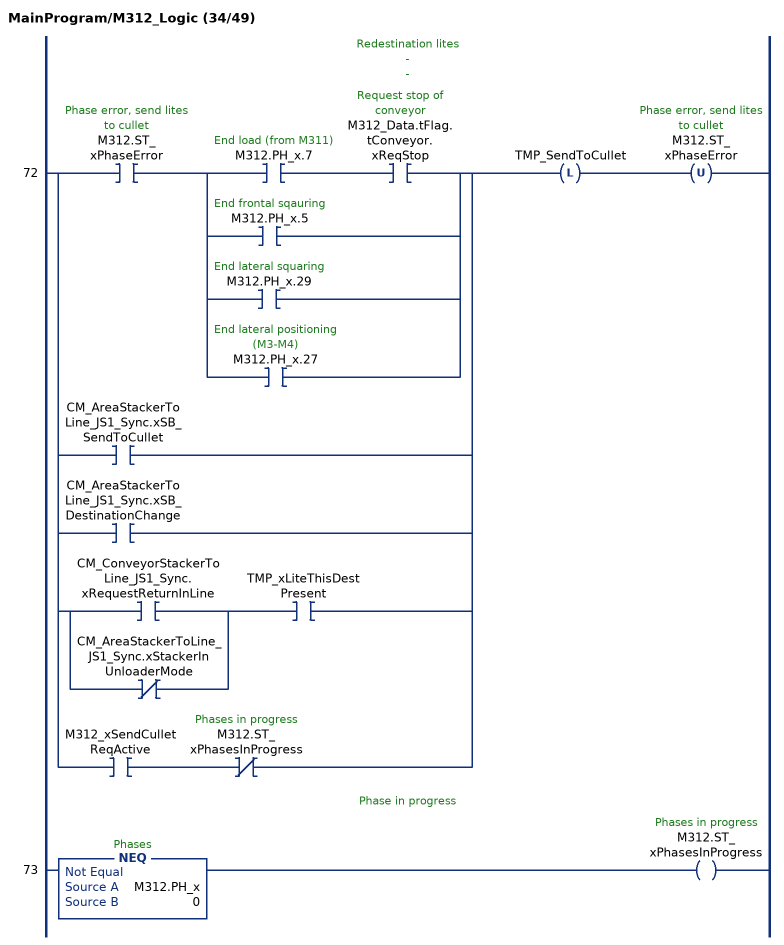
   // Redestination lites
   // -
   // -
   72: [XIC(M312.ST_xPhaseError) [XIC(M312.PH_x.7) XIC(M312_Data.tFlag.tConveyor.xReqStop) ,XIC(M312.PH_x.5) ,XIC(M312.PH_x.29) ,XIC(M312.PH_x.27) ] ,[XIC(CM_AreaStackerToLine_JS1_Sync.xSB_SendToCullet) ,XIC(CM_AreaStackerToLine_JS1_Sync.xSB_DestinationChange) ] ,[XIC(CM_ConveyorStackerToLine_JS1_Sync.xRequestReturnInLine) ,XIO(CM_AreaStackerToLine_JS1_Sync.xStackerInUnloaderMode) ] XIC(TMP_xLiteThisDestPresent) ,XIC(M312_xSendCulletReqActive) XIO(M312.ST_xPhasesInProgress) ]OTL(TMP_SendToCullet)OTU(M312.ST_xPhaseError);
   // Phase in progress
   73: NEQ(M312.PH_x,0)OTE(M312.ST_xPhasesInProgress);
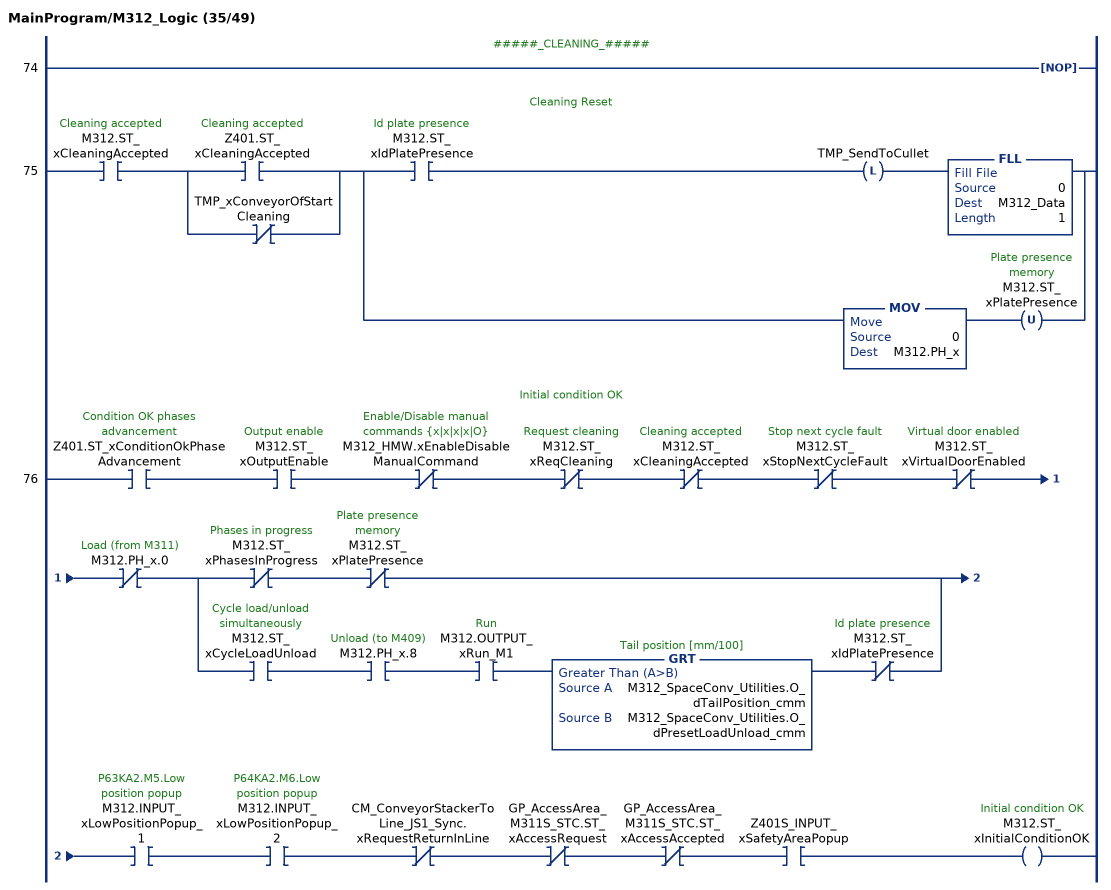
   // #####_CLEANING_#####
   74: NOP();
   // Cleaning Reset
   75: XIC(M312.ST_xCleaningAccepted)[XIC(Z401.ST_xCleaningAccepted) ,XIO(TMP_xConveyorOfStartCleaning) ][XIC(M312.ST_xIdPlatePresence) OTL(TMP_SendToCullet) FLL(0,M312_Data,1) ,MOV(0,M312.PH_x) OTU(M312.ST_xPlatePresence) ];
   // Initial condition OK
   76: XIC(Z401.ST_xConditionOkPhaseAdvancement)XIC(M312.ST_xOutputEnable)XIO(M312_HMW.xEnableDisableManualCommand)XIO(M312.ST_xReqCleaning)XIO(M312.ST_xCleaningAccepted)XIO(M312.ST_xStopNextCycleFault)XIO(M312.ST_xVirtualDoorEnabled)XIO(M312.PH_x.0)[XIO(M312.ST_xPhasesInProgress) XIO(M312.ST_xPlatePresence) ,XIC(M312.ST_xCycleLoadUnload) XIC(M312.PH_x.8) XIC(M312.OUTPUT_xRun_M1) GRT(M312_SpaceConv_Utilities.O_dTailPosition_cmm,M312_SpaceConv_Utilities.O_dPresetLoadUnload_cmm) XIO(M312.ST_xIdPlatePresence) ]XIC(M312.INPUT_xLowPositionPopup_1)XIC(M312.INPUT_xLowPositionPopup_2)XIO(CM_ConveyorStackerToLine_JS1_Sync.xRequestReturnInLine)XIO(GP_AccessArea_M311S_STC.ST_xAccessRequest)XIO(GP_AccessArea_M311S_STC.ST_xAccessAccepted)XIC(Z401S_INPUT_xSafetyAreaPopup)OTE(M312.ST_xInitialConditionOK);
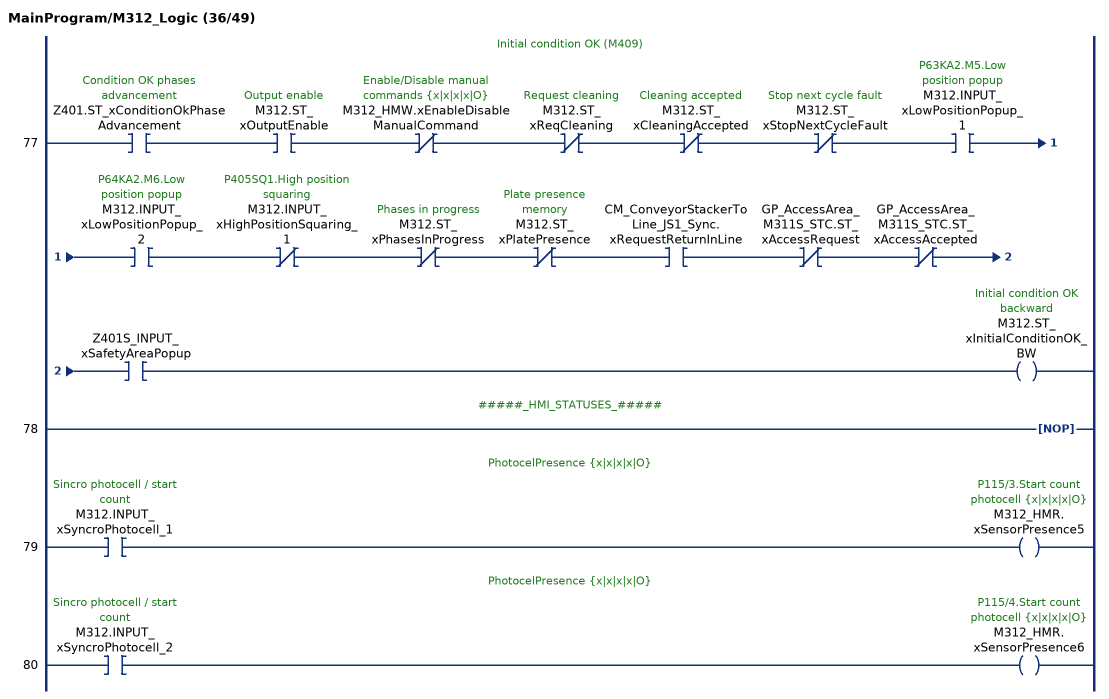
   // Initial condition OK (M409)
   77: XIC(Z401.ST_xConditionOkPhaseAdvancement)XIC(M312.ST_xOutputEnable)XIO(M312_HMW.xEnableDisableManualCommand)XIO(M312.ST_xReqCleaning)XIO(M312.ST_xCleaningAccepted)XIO(M312.ST_xStopNextCycleFault)XIC(M312.INPUT_xLowPositionPopup_1)XIC(M312.INPUT_xLowPositionPopup_2)XIO(M312.INPUT_xHighPositionSquaring_1)XIO(M312.ST_xPhasesInProgress)XIO(M312.ST_xPlatePresence)XIC(CM_ConveyorStackerToLine_JS1_Sync.xRequestReturnInLine)XIO(GP_AccessArea_M311S_STC.ST_xAccessRequest)XIO(GP_AccessArea_M311S_STC.ST_xAccessAccepted)XIC(Z401S_INPUT_xSafetyAreaPopup)OTE(M312.ST_xInitialConditionOK_BW);
   // #####_HMI_STATUSES_#####
   78: NOP();
   // PhotocelPresence {x|x|x|x|O}
   79: XIC(M312.INPUT_xSyncroPhotocell_1)OTE(M312_HMR.xSensorPresence5);
   // PhotocelPresence {x|x|x|x|O}
   80: XIC(M312.INPUT_xSyncroPhotocell_2)OTE(M312_HMR.xSensorPresence6);
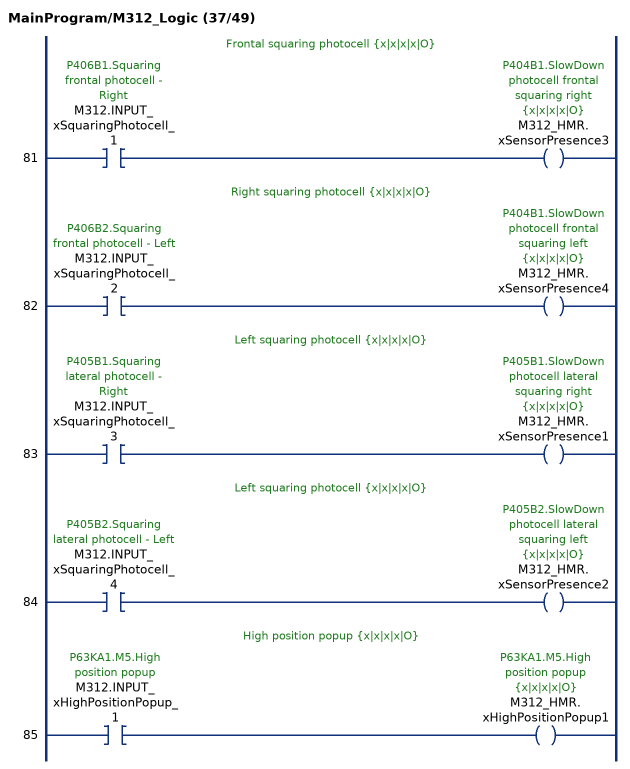
   // Frontal squaring photocell {x|x|x|x|O}
   81: XIC(M312.INPUT_xSquaringPhotocell_1)OTE(M312_HMR.xSensorPresence3);
   // Right squaring photocell {x|x|x|x|O}
   82: XIC(M312.INPUT_xSquaringPhotocell_2)OTE(M312_HMR.xSensorPresence4);
   // Left squaring photocell {x|x|x|x|O}
   83: XIC(M312.INPUT_xSquaringPhotocell_3)OTE(M312_HMR.xSensorPresence1);
   // Left squaring photocell {x|x|x|x|O}
   84: XIC(M312.INPUT_xSquaringPhotocell_4)OTE(M312_HMR.xSensorPresence2);
   // High position popup {x|x|x|x|O}
   85: XIC(M312.INPUT_xHighPositionPopup_1)OTE(M312_HMR.xHighPositionPopup1);
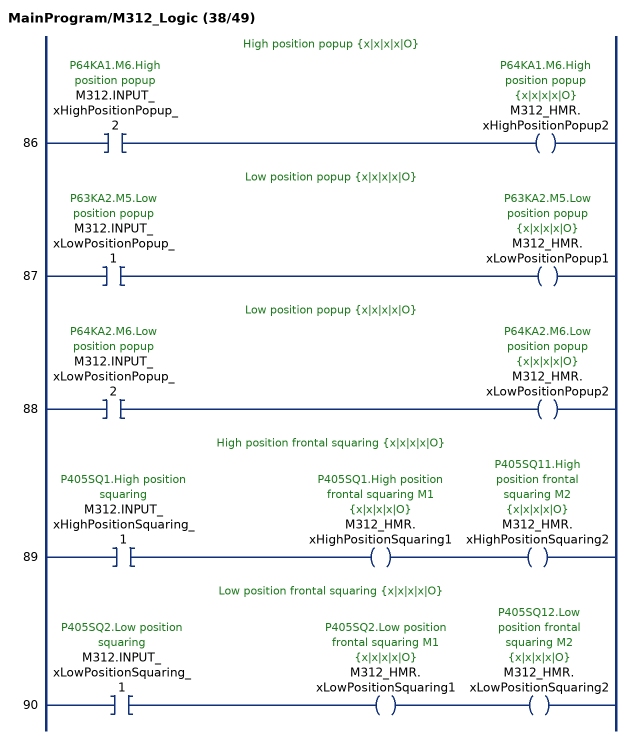
   // High position popup {x|x|x|x|O}
   86: XIC(M312.INPUT_xHighPositionPopup_2)OTE(M312_HMR.xHighPositionPopup2);
   // Low position popup {x|x|x|x|O}
   87: XIC(M312.INPUT_xLowPositionPopup_1)OTE(M312_HMR.xLowPositionPopup1);
   // Low position popup {x|x|x|x|O}
   88: XIC(M312.INPUT_xLowPositionPopup_2)OTE(M312_HMR.xLowPositionPopup2);
   // High position frontal squaring {x|x|x|x|O}
   89: XIC(M312.INPUT_xHighPositionSquaring_1)OTE(M312_HMR.xHighPositionSquaring1)OTE(M312_HMR.xHighPositionSquaring2);
   // Low position frontal squaring {x|x|x|x|O}
   90: XIC(M312.INPUT_xLowPositionSquaring_1)OTE(M312_HMR.xLowPositionSquaring1)OTE(M312_HMR.xLowPositionSquaring2);
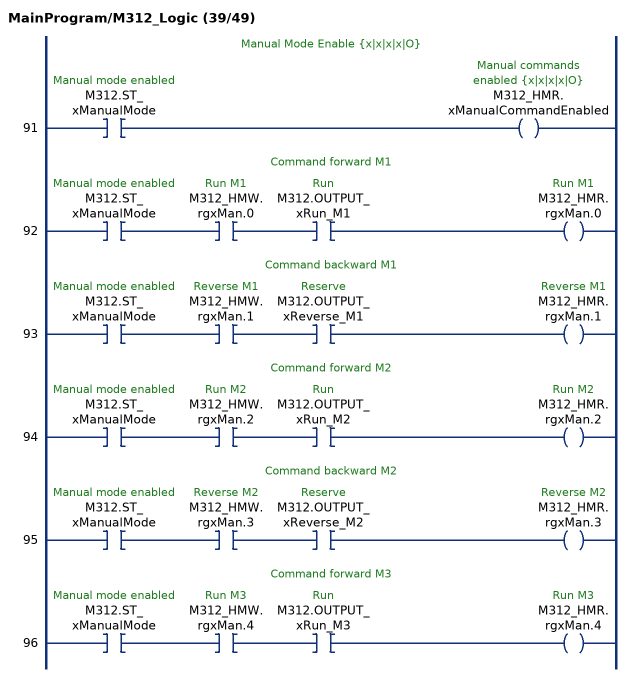
   // Manual Mode Enable {x|x|x|x|O}
   91: XIC(M312.ST_xManualMode)OTE(M312_HMR.xManualCommandEnabled);
   // Command forward M1
   92: XIC(M312.ST_xManualMode)XIC(M312_HMW.rgxMan.0)XIC(M312.OUTPUT_xRun_M1)OTE(M312_HMR.rgxMan.0);
   // Command backward M1
   93: XIC(M312.ST_xManualMode)XIC(M312_HMW.rgxMan.1)XIC(M312.OUTPUT_xReverse_M1)OTE(M312_HMR.rgxMan.1);
   // Command forward M2
   94: XIC(M312.ST_xManualMode)XIC(M312_HMW.rgxMan.2)XIC(M312.OUTPUT_xRun_M2)OTE(M312_HMR.rgxMan.2);
   // Command backward M2
   95: XIC(M312.ST_xManualMode)XIC(M312_HMW.rgxMan.3)XIC(M312.OUTPUT_xReverse_M2)OTE(M312_HMR.rgxMan.3);
   // Command forward M3
   96: XIC(M312.ST_xManualMode)XIC(M312_HMW.rgxMan.4)XIC(M312.OUTPUT_xRun_M3)OTE(M312_HMR.rgxMan.4);
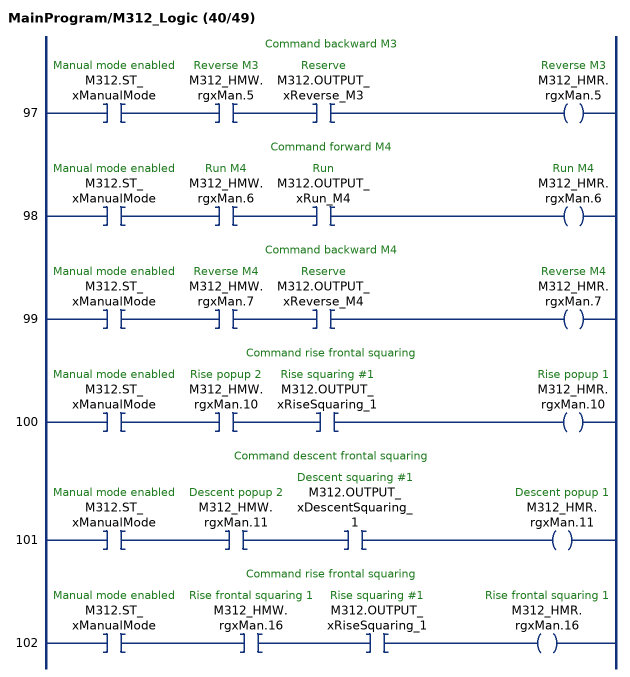
   // Command backward M3
   97: XIC(M312.ST_xManualMode)XIC(M312_HMW.rgxMan.5)XIC(M312.OUTPUT_xReverse_M3)OTE(M312_HMR.rgxMan.5);
   // Command forward M4
   98: XIC(M312.ST_xManualMode)XIC(M312_HMW.rgxMan.6)XIC(M312.OUTPUT_xRun_M4)OTE(M312_HMR.rgxMan.6);
   // Command backward M4
   99: XIC(M312.ST_xManualMode)XIC(M312_HMW.rgxMan.7)XIC(M312.OUTPUT_xReverse_M4)OTE(M312_HMR.rgxMan.7);
   // Command rise frontal squaring
   100: XIC(M312.ST_xManualMode)XIC(M312_HMW.rgxMan.10)XIC(M312.OUTPUT_xRiseSquaring_1)OTE(M312_HMR.rgxMan.10);
   // Command descent frontal squaring
   101: XIC(M312.ST_xManualMode)XIC(M312_HMW.rgxMan.11)XIC(M312.OUTPUT_xDescentSquaring_1)OTE(M312_HMR.rgxMan.11);
   // Command rise frontal squaring
   102: XIC(M312.ST_xManualMode)XIC(M312_HMW.rgxMan.16)XIC(M312.OUTPUT_xRiseSquaring_1)OTE(M312_HMR.rgxMan.16);
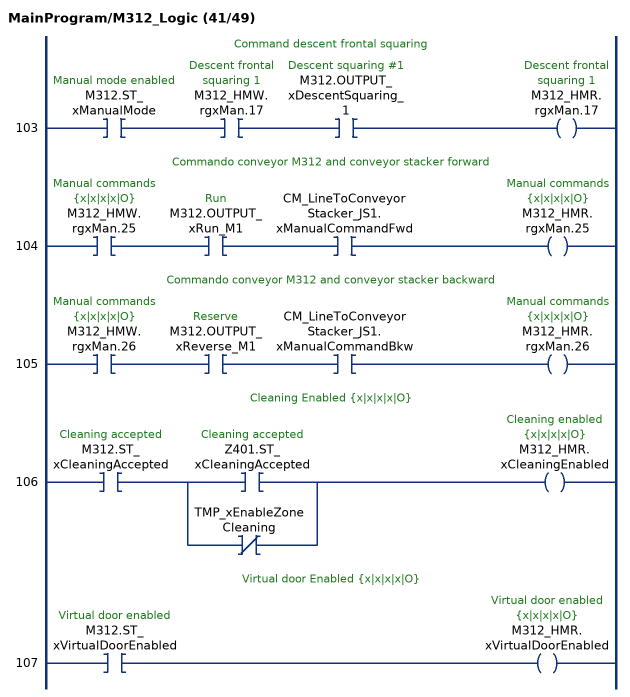
   // Command descent frontal squaring
   103: XIC(M312.ST_xManualMode)XIC(M312_HMW.rgxMan.17)XIC(M312.OUTPUT_xDescentSquaring_1)OTE(M312_HMR.rgxMan.17);
   // Commando conveyor M312 and conveyor stacker forward
   104: XIC(M312_HMW.rgxMan.25)XIC(M312.OUTPUT_xRun_M1)XIC(CM_LineToConveyorStacker_JS1.xManualCommandFwd)OTE(M312_HMR.rgxMan.25);
   // Commando conveyor M312 and conveyor stacker backward
   105: XIC(M312_HMW.rgxMan.26)XIC(M312.OUTPUT_xReverse_M1)XIC(CM_LineToConveyorStacker_JS1.xManualCommandBkw)OTE(M312_HMR.rgxMan.26);
   // Cleaning Enabled {x|x|x|x|O}
   106: XIC(M312.ST_xCleaningAccepted)[XIC(Z401.ST_xCleaningAccepted) ,XIO(TMP_xEnableZoneCleaning) ]OTE(M312_HMR.xCleaningEnabled);
   // Virtual door Enabled {x|x|x|x|O}
   107: XIC(M312.ST_xVirtualDoorEnabled)OTE(M312_HMR.xVirtualDoorEnabled);
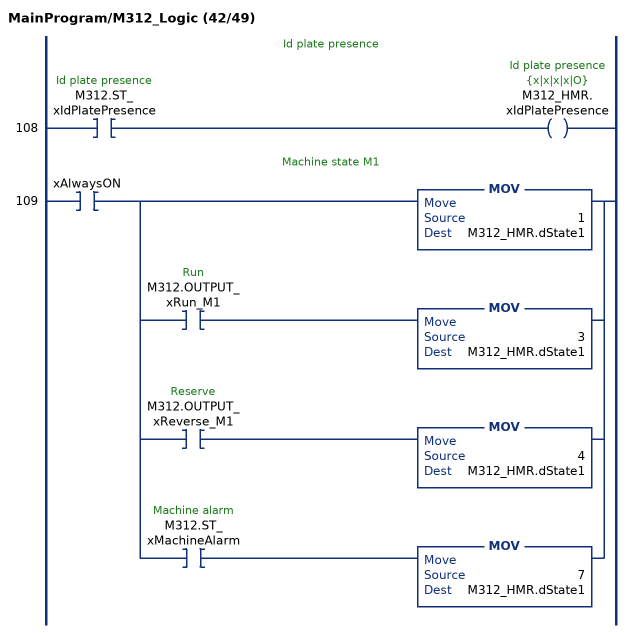
   // Id plate presence
   108: XIC(M312.ST_xIdPlatePresence)OTE(M312_HMR.xIdPlatePresence);
   // Machine state M1
   109: XIC(xAlwaysON)[MOV(1,M312_HMR.dState1) ,XIC(M312.OUTPUT_xRun_M1) MOV(3,M312_HMR.dState1) ,XIC(M312.OUTPUT_xReverse_M1) MOV(4,M312_HMR.dState1) ,XIC(M312.ST_xMachineAlarm) MOV(7,M312_HMR.dState1) ];
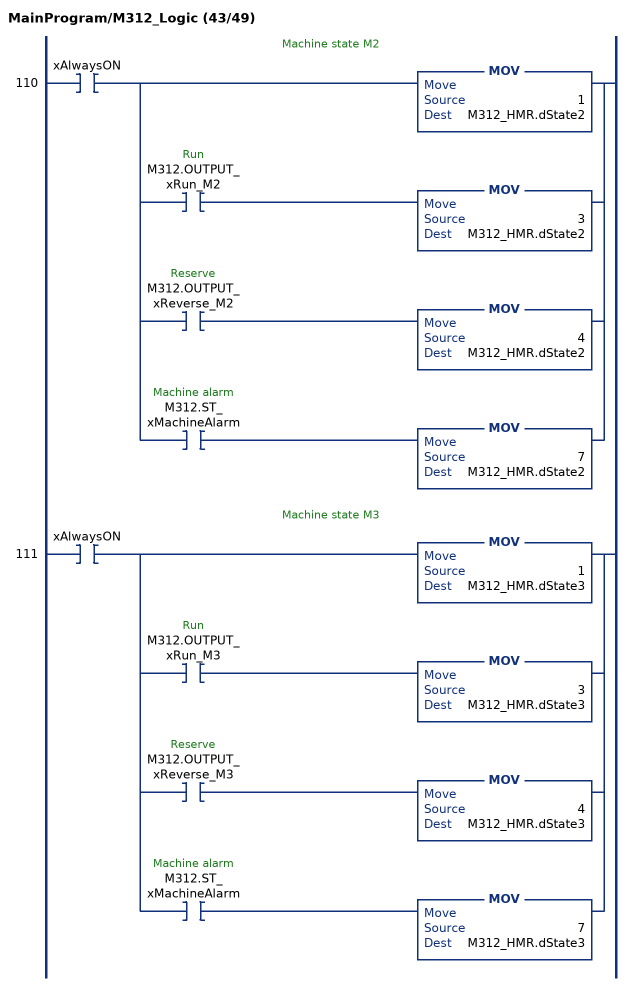
   // Machine state M2
   110: XIC(xAlwaysON)[MOV(1,M312_HMR.dState2) ,XIC(M312.OUTPUT_xRun_M2) MOV(3,M312_HMR.dState2) ,XIC(M312.OUTPUT_xReverse_M2) MOV(4,M312_HMR.dState2) ,XIC(M312.ST_xMachineAlarm) MOV(7,M312_HMR.dState2) ];
   // Machine state M3
   111: XIC(xAlwaysON)[MOV(1,M312_HMR.dState3) ,XIC(M312.OUTPUT_xRun_M3) MOV(3,M312_HMR.dState3) ,XIC(M312.OUTPUT_xReverse_M3) MOV(4,M312_HMR.dState3) ,XIC(M312.ST_xMachineAlarm) MOV(7,M312_HMR.dState3) ];
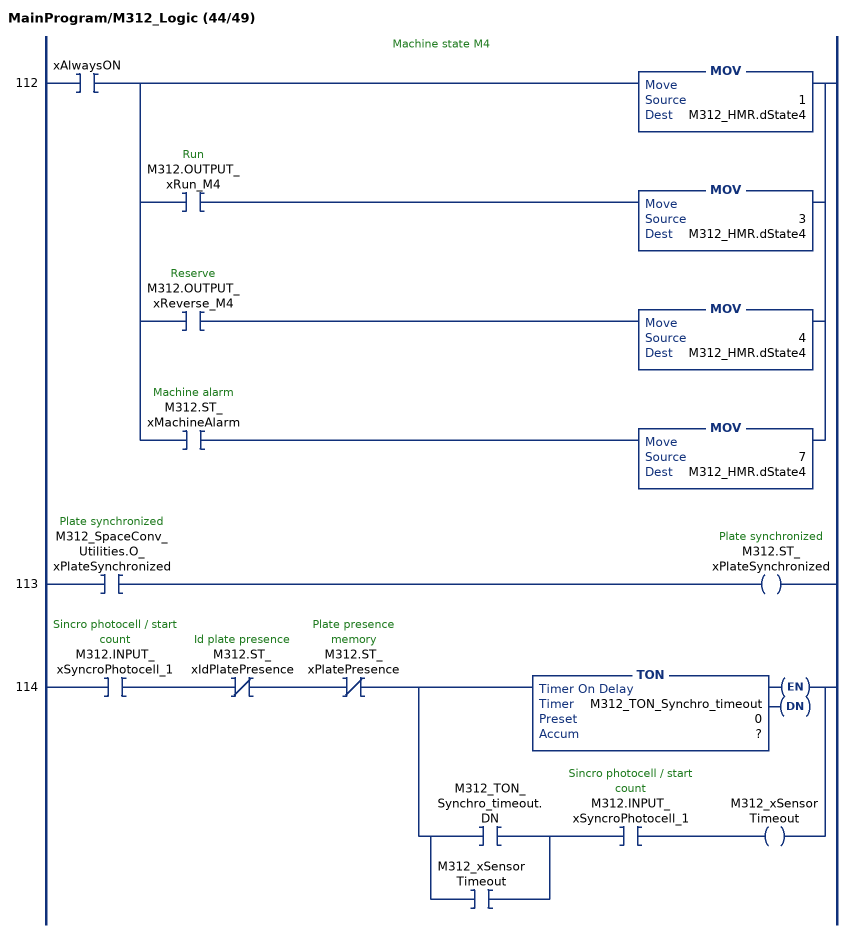
   // Machine state M4
   112: XIC(xAlwaysON)[MOV(1,M312_HMR.dState4) ,XIC(M312.OUTPUT_xRun_M4) MOV(3,M312_HMR.dState4) ,XIC(M312.OUTPUT_xReverse_M4) MOV(4,M312_HMR.dState4) ,XIC(M312.ST_xMachineAlarm) MOV(7,M312_HMR.dState4) ];
   113: XIC(M312_SpaceConv_Utilities.O_xPlateSynchronized)OTE(M312.ST_xPlateSynchronized);
   114: XIC(M312.INPUT_xSyncroPhotocell_1)XIO(M312.ST_xIdPlatePresence)XIO(M312.ST_xPlatePresence)[TON(M312_TON_Synchro_timeout,?,?) ,[XIC(M312_TON_Synchro_timeout.DN) ,XIC(M312_xSensorTimeout) ] XIC(M312.INPUT_xSyncroPhotocell_1) OTE(M312_xSensorTimeout) ];
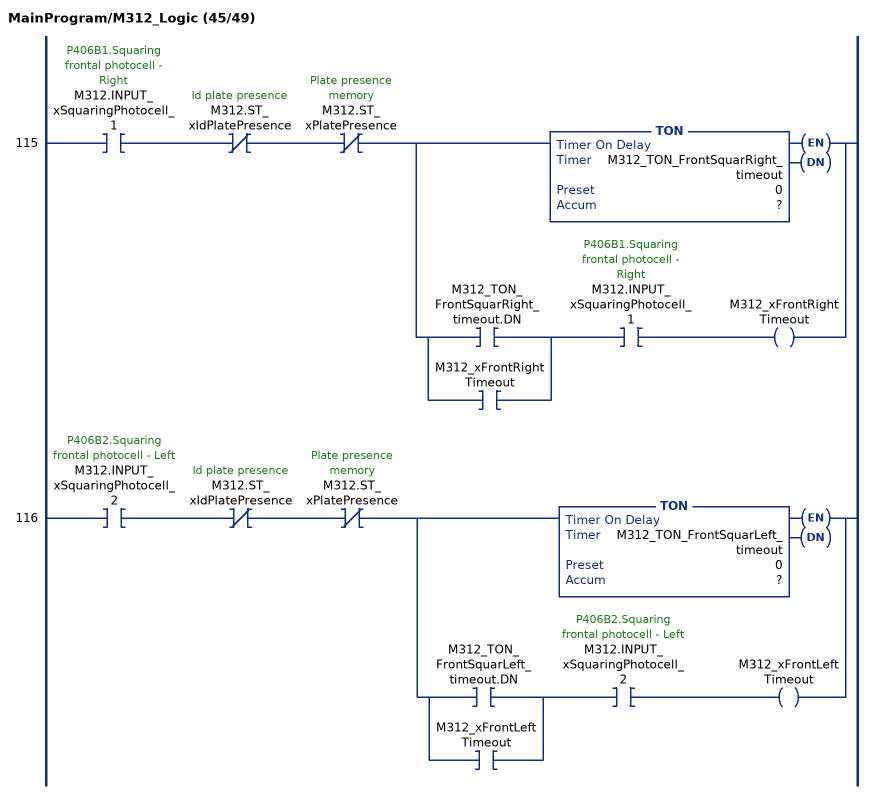
   115: XIC(M312.INPUT_xSquaringPhotocell_1)XIO(M312.ST_xIdPlatePresence)XIO(M312.ST_xPlatePresence)[TON(M312_TON_FrontSquarRight_timeout,?,?) ,[XIC(M312_TON_FrontSquarRight_timeout.DN) ,XIC(M312_xFrontRightTimeout) ] XIC(M312.INPUT_xSquaringPhotocell_1) OTE(M312_xFrontRightTimeout) ];
   116: XIC(M312.INPUT_xSquaringPhotocell_2)XIO(M312.ST_xIdPlatePresence)XIO(M312.ST_xPlatePresence)[TON(M312_TON_FrontSquarLeft_timeout,?,?) ,[XIC(M312_TON_FrontSquarLeft_timeout.DN) ,XIC(M312_xFrontLeftTimeout) ] XIC(M312.INPUT_xSquaringPhotocell_2) OTE(M312_xFrontLeftTimeout) ];
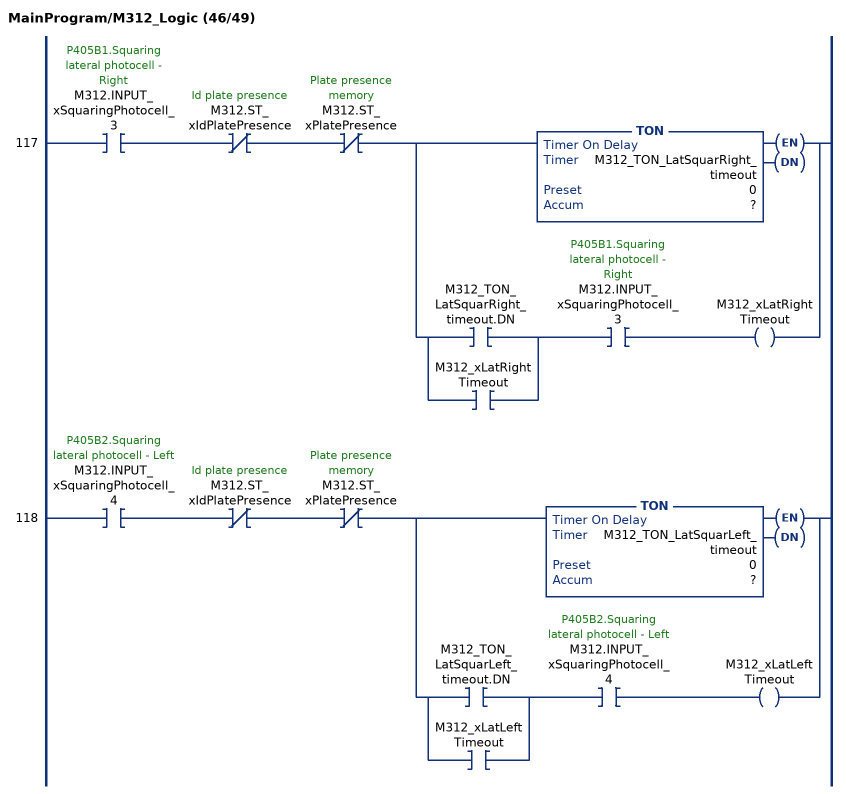
   117: XIC(M312.INPUT_xSquaringPhotocell_3)XIO(M312.ST_xIdPlatePresence)XIO(M312.ST_xPlatePresence)[TON(M312_TON_LatSquarRight_timeout,?,?) ,[XIC(M312_TON_LatSquarRight_timeout.DN) ,XIC(M312_xLatRightTimeout) ] XIC(M312.INPUT_xSquaringPhotocell_3) OTE(M312_xLatRightTimeout) ];
   118: XIC(M312.INPUT_xSquaringPhotocell_4)XIO(M312.ST_xIdPlatePresence)XIO(M312.ST_xPlatePresence)[TON(M312_TON_LatSquarLeft_timeout,?,?) ,[XIC(M312_TON_LatSquarLeft_timeout.DN) ,XIC(M312_xLatLeftTimeout) ] XIC(M312.INPUT_xSquaringPhotocell_4) OTE(M312_xLatLeftTimeout) ];
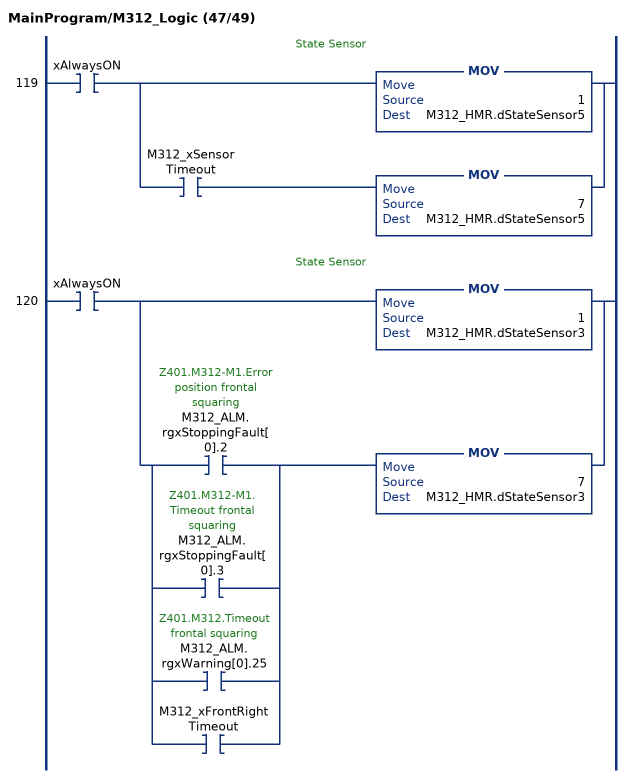
   // State Sensor
   119: XIC(xAlwaysON)[MOV(1,M312_HMR.dStateSensor5) ,XIC(M312_xSensorTimeout) MOV(7,M312_HMR.dStateSensor5) ];
   // State Sensor
   120: XIC(xAlwaysON)[MOV(1,M312_HMR.dStateSensor3) ,[XIC(M312_ALM.rgxStoppingFault[0].2) ,XIC(M312_ALM.rgxStoppingFault[0].3) ,XIC(M312_ALM.rgxWarning[0].25) ,XIC(M312_xFrontRightTimeout) ] MOV(7,M312_HMR.dStateSensor3) ];
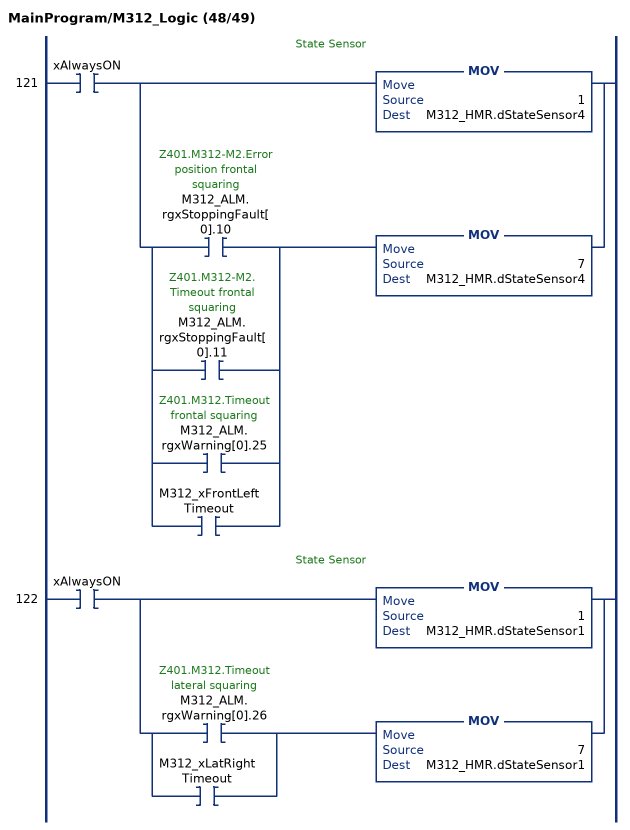
   // State Sensor
   121: XIC(xAlwaysON)[MOV(1,M312_HMR.dStateSensor4) ,[XIC(M312_ALM.rgxStoppingFault[0].10) ,XIC(M312_ALM.rgxStoppingFault[0].11) ,XIC(M312_ALM.rgxWarning[0].25) ,XIC(M312_xFrontLeftTimeout) ] MOV(7,M312_HMR.dStateSensor4) ];
   // State Sensor
   122: XIC(xAlwaysON)[MOV(1,M312_HMR.dStateSensor1) ,[XIC(M312_ALM.rgxWarning[0].26) ,XIC(M312_xLatRightTimeout) ] MOV(7,M312_HMR.dStateSensor1) ];
